// TIA Portal project "Proyecto_final" (V15.1)

(* hardware
DEVICE "S71500/ET200MP station_1"  S7-1500 station
   slot 0: "Rail_0"  Rack  6ES7 590-1***0-0AA0
   slot 1: "PLC_1"  CPU 1516-3 PN/DP  6ES7 516-3AN01-0AB0  V2.6
      slot 3: "CPU display_1"  6ES7591-1BA00-0AA0
   slot 2: "AI 8xU/I/RTD/TC ST_1"  AI 8xU/I/RTD/TC ST  6ES7 531-7KF00-0AB0  V2.2
   slot 3: "AQ 4xU/I ST_1"  AQ 4xU/I ST  6ES7 532-5HD00-0AB0  V2.2
   slot 4: "DI 32x24VDC HF_1"  DI 32x24VDC HF  6ES7 521-1BL00-0AB0  V2.1
   slot 5: "DQ 32x24VDC/0.5A HF_1"  DQ 32x24VDC/0.5A HF  6ES7 522-1BL01-0AB0  V1.1
DEVICE "S7-1200 station_1"  S7-1200 Station
   slot 0: "Rack_0"  S7-1200 Rack  Rack  V1.0
   slot 1: "PLC_2"  CPU 1215C DC/DC/DC  6ES7 215-1AG40-0XB0  V4.2
DEVICE "S7-1200 station_2"  S7-1200 Station
   slot 0: "Rack_0"  S7-1200 Rack  Rack  V1.0
   slot 1: "PLC_3"  CPU 1215C DC/DC/DC  6ES7 215-1AG40-0XB0  V4.2
DEVICE "HMI_1"  KTP400 Basic PN
   slot 0: "HMI_1"  KTP400 Basic PN  6AV2 123-2DB03-0AX0  15.1.0.0
   slot 1: "HMI_RT_1"  KTP400 Basic PN  6AV2 123-2DB03-0AX0  15.1.0.0
   slot 5: "HMI_1.IE_CP_1"  PROFINET Interface  15.0.1.0
      slot 1: "PROFINET Interface_1"  PROFINET Interface
         slot 1: "Port_1"  Port
DEVICE "HMI_2"  KTP400 Basic PN
   slot 0: "HMI_2"  KTP400 Basic PN  6AV2 123-2DB03-0AX0  15.1.0.0
   slot 1: "HMI_RT_2"  KTP400 Basic PN  6AV2 123-2DB03-0AX0  15.1.0.0
   slot 5: "HMI_2.IE_CP_1"  PROFINET Interface  15.0.1.0
      slot 1: "PROFINET Interface_1"  PROFINET Interface
         slot 1: "Port_1"  Port
DEVICE "HMI_3"  KTP400 Basic PN
   slot 0: "HMI_3"  KTP400 Basic PN  6AV2 123-2DB03-0AX0  15.1.0.0
   slot 1: "HMI_RT_3"  KTP400 Basic PN  6AV2 123-2DB03-0AX0  15.1.0.0
   slot 5: "HMI_3.IE_CP_1"  PROFINET Interface  15.0.1.0
      slot 1: "PROFINET Interface_1"  PROFINET Interface
         slot 1: "Port_1"  Port
DEVICE "SCALANCE X005"  SCALANCE X-Station
   slot 0: "SCALANCE X rack"  Rail
   slot 0: "Switch_1"  6GK5 005-0BA00-1AB2  V1.0
*)

// ===== PLC "PLC_1"  CPU 1516-3 PN/DP =====

VAR_GLOBAL   // PLC tag table "Default tag table"
   "Encendido" AT %M8.0 : Bool;
   "PE" AT %I17.3 : Bool;
   "Tag_1" AT %Q9.3 : Bool;
   "Tag_2" AT %Q9.4 : Bool;
   "LED_estado" AT %Q9.5 : Bool;
   "LED_PE" AT %Q9.6 : Bool;
   "Tag_3" AT %I17.4 : Bool;
   "Tag_4" AT %I17.5 : Bool;
   "Tag_5" AT %I17.6 : Bool;
END_VAR

DATA_BLOCK "PLC1_Ban"   // DB2
{ S7_Optimized_Access := 'FALSE' }
VERSION : 0.1
   VAR
      Ban_estado : Bool;
      Ban_dirección : UInt;
   END_VAR
BEGIN
END_DATA_BLOCK

// folder: System blocks/Program resources

DATA_BLOCK "IEC_Timer_0_DB"   // DB1
{ S7_Optimized_Access := 'TRUE' }
AUTHOR : Simatic
FAMILY : IEC
NAME : IEC_TMR
VERSION : 1.0
// stored: InstanceOfName IEC_TIMER
"IEC_TIMER"
BEGIN
END_DATA_BLOCK

// folder: (top level)

ORGANIZATION_BLOCK "Main"   // OB1, LAD, ProgramCycle
TITLE = Control de banda transportadora
{ S7_Optimized_Access := 'TRUE' }
VERSION : 0.1
   VAR_INPUT
      Initial_Call : Bool;   // Initial call of this OB
      Remanence : Bool;   // =True, if remanent data are available
   END_VAR
   VAR_TEMP   // added for the SCL form of the ladder/FBD networks
      _w1 : Bool;
   END_VAR
BEGIN

REGION Network 1: Control motor
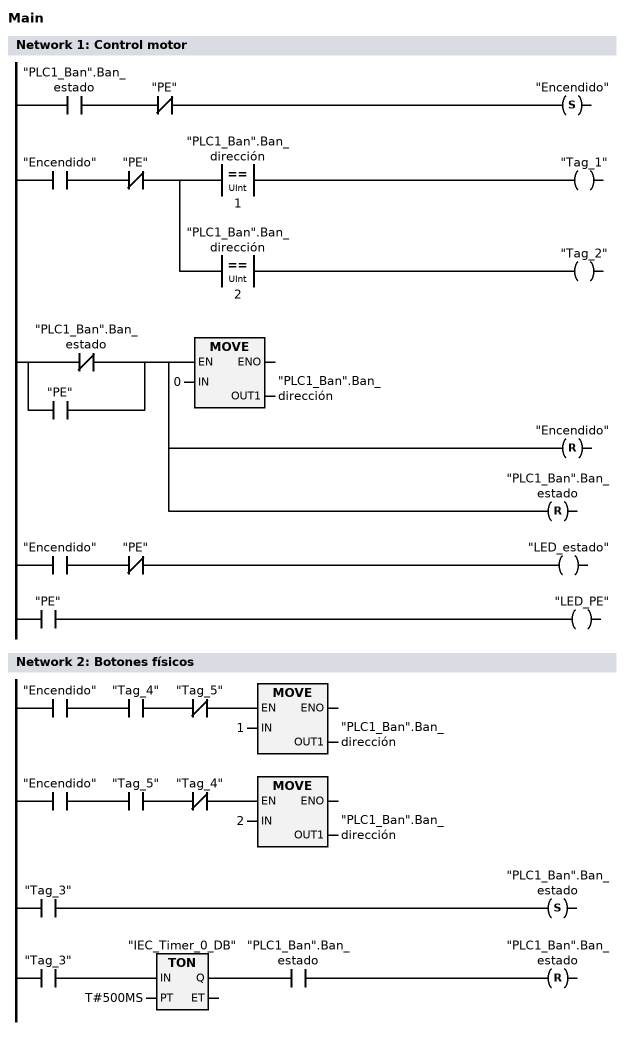
   RUNG wire#powerrail
      Contact( "PLC1_Ban".Ban_estado )
      I_Contact( "PE" )
      S_Coil( "Encendido" )
   END_RUNG
   RUNG wire#powerrail
      Contact( "Encendido" )
      I_Contact( "PE" )
      wire#w1
      { S7_Templates := "SrcType := UInt" } EQ_Contact(in1 := "PLC1_Ban".Ban_dirección, in2 := 1)
      Coil( "Tag_1" )
   END_RUNG
   RUNG wire#w1
      { S7_Templates := "SrcType := UInt" } EQ_Contact(in1 := "PLC1_Ban".Ban_dirección, in2 := 2)
      Coil( "Tag_2" )
   END_RUNG
   RUNG wire#powerrail
      I_Contact( "PLC1_Ban".Ban_estado )
      wire#w2
      Move(in := 0, out1 => "PLC1_Ban".Ban_dirección)
   END_RUNG
   RUNG wire#powerrail
      Contact( "PE" )
   END_RUNG wire#w2
   RUNG wire#w2
      R_Coil( "Encendido" )
   END_RUNG
   RUNG wire#w2
      R_Coil( "PLC1_Ban".Ban_estado )
   END_RUNG
   RUNG wire#powerrail
      Contact( "Encendido" )
      I_Contact( "PE" )
      Coil( "LED_estado" )
   END_RUNG
   RUNG wire#powerrail
      Contact( "PE" )
      Coil( "LED_PE" )
   END_RUNG
   // the same network as SCL:
   IF "PLC1_Ban".Ban_estado AND NOT "PE" THEN "Encendido" := TRUE; END_IF;
   #_w1 := "Encendido" AND NOT "PE";
   "Tag_1" := #_w1 AND ("PLC1_Ban".Ban_dirección = 1);
   "Tag_2" := #_w1 AND ("PLC1_Ban".Ban_dirección = 2);
   IF NOT "PLC1_Ban".Ban_estado OR "PE" THEN
       "PLC1_Ban".Ban_dirección := 0;
       "Encendido" := FALSE;
       "PLC1_Ban".Ban_estado := FALSE;
   END_IF;
   "LED_estado" := "Encendido" AND NOT "PE";
   "LED_PE" := "PE";
END_REGION

REGION Network 2: Botones físicos
   IF "Encendido" AND "Tag_4" AND NOT "Tag_5" THEN "PLC1_Ban".Ban_dirección := 1; END_IF;
   IF "Encendido" AND "Tag_5" AND NOT "Tag_4" THEN "PLC1_Ban".Ban_dirección := 2; END_IF;
   IF "Tag_3" THEN "PLC1_Ban".Ban_estado := TRUE; END_IF;
   "IEC_Timer_0_DB".TON(IN := "Tag_3", PT := T#500MS);
   IF "IEC_Timer_0_DB".Q AND "PLC1_Ban".Ban_estado THEN "PLC1_Ban".Ban_estado := FALSE; END_IF;
END_REGION
END_ORGANIZATION_BLOCK

// ===== PLC "PLC_2"  CPU 1215C DC/DC/DC =====

VAR_GLOBAL   // PLC tag table "Default tag table"
   "Rev_Detección" AT %M0.1 : Bool;
   "Rev_especial" AT %MW4 : UInt;
   "Rev_estado" AT %M0.0 : Bool;
   "Rev_progreso" AT %MW2 : Int;
   "B4" AT %I0.0 : Bool;
   "F3" AT %Q0.0 : Bool;
   "F2" AT %Q0.1 : Bool;
   "F1" AT %Q0.2 : Bool;
   "Piston_arriba" AT %Q0.3 : Bool;
   "Piston_abajo" AT %Q0.4 : Bool;
   "PE" AT %I0.4 : Bool;
   "Sens_abajo" AT %I0.5 : Bool;
   "Sens_arriba" AT %I0.6 : Bool;
   "B3" AT %I0.1 : Bool;
   "B2" AT %I0.2 : Bool;
   "B1" AT %I0.3 : Bool;
   "Encendido" AT %M0.2 : Bool;
   "Fin" AT %M0.3 : Bool;
   "Ciclo" AT %M0.4 : Bool;
   "Mem_pos" AT %M0.5 : Bool;
   "Cuenta_add" AT %MW6 : Int;
   "Reset" AT %M0.6 : Bool;
   "Skip" AT %M0.7 : Bool;
   "Tag_1" AT %M8.0 : Bool;
END_VAR

DATA_BLOCK "PLC2_Rev"   // DB5
{ S7_Optimized_Access := 'FALSE' }
VERSION : 0.1
   VAR
      Rev_Detección : Bool;
      Rev_especial : UInt;
      Rev_estado : Bool;
      Rev_progreso : Int;
   END_VAR
BEGIN
END_DATA_BLOCK

// folder: System blocks/Program resources

DATA_BLOCK "IEC_Timer_0_DB"   // DB1
{ S7_Optimized_Access := 'TRUE' }
AUTHOR : Simatic
FAMILY : IEC
NAME : IEC_TMR
VERSION : 1.0
// stored: InstanceOfName IEC_TIMER
"IEC_TIMER"
BEGIN
END_DATA_BLOCK

DATA_BLOCK "IEC_Counter_0_DB"   // DB2
{ S7_Optimized_Access := 'TRUE' }
AUTHOR : Simatic
FAMILY : IEC
NAME : CNTR
VERSION : 1.0
// stored: InstanceOfName IEC_COUNTER
"IEC_COUNTER"
BEGIN
END_DATA_BLOCK

DATA_BLOCK "IEC_Timer_0_DB_2"   // DB3
{ S7_Optimized_Access := 'TRUE' }
AUTHOR : Simatic
FAMILY : IEC
NAME : IEC_TMR
VERSION : 1.0
// stored: InstanceOfName IEC_TIMER
"IEC_TIMER"
BEGIN
END_DATA_BLOCK

DATA_BLOCK "IEC_Timer_0_DB_1"   // DB4
{ S7_Optimized_Access := 'TRUE' }
AUTHOR : Simatic
FAMILY : IEC
NAME : IEC_TMR
VERSION : 1.0
// stored: InstanceOfName IEC_TIMER
"IEC_TIMER"
BEGIN
END_DATA_BLOCK

DATA_BLOCK "IEC_Timer_0_DB_3"   // DB6
{ S7_Optimized_Access := 'TRUE' }
AUTHOR : Simatic
FAMILY : IEC
NAME : IEC_TMR
VERSION : 1.0
// stored: InstanceOfName IEC_TIMER
"IEC_TIMER"
BEGIN
END_DATA_BLOCK

DATA_BLOCK "IEC_Timer_0_DB_4"   // DB7
{ S7_Optimized_Access := 'TRUE' }
AUTHOR : Simatic
FAMILY : IEC
NAME : IEC_TMR
VERSION : 1.0
// stored: InstanceOfName IEC_TIMER
"IEC_TIMER"
BEGIN
END_DATA_BLOCK

DATA_BLOCK "IEC_Timer_0_DB_5"   // DB8
{ S7_Optimized_Access := 'TRUE' }
AUTHOR : Simatic
FAMILY : IEC
NAME : IEC_TMR
VERSION : 1.0
// stored: InstanceOfName IEC_TIMER
"IEC_TIMER"
BEGIN
END_DATA_BLOCK

// folder: (top level)

ORGANIZATION_BLOCK "Main"   // OB1, LAD, ProgramCycle
TITLE = Revolvedora
{ S7_Optimized_Access := 'TRUE' }
VERSION : 0.1
   VAR_INPUT
      Initial_Call : Bool;   // Initial call of this OB
      Remanence : Bool;   // =True, if remanent data are available
   END_VAR
   VAR_TEMP   // added for the SCL form of the ladder/FBD networks
      _w1 : Bool;
   END_VAR
BEGIN

REGION Network 1
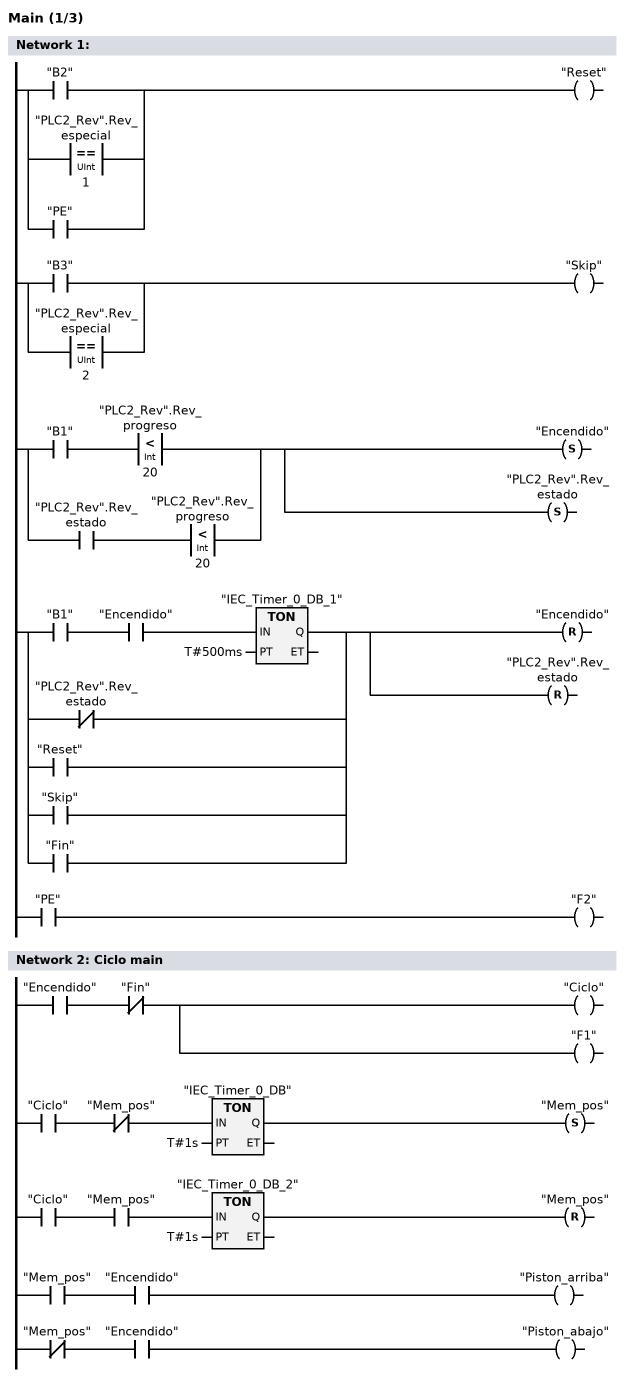
   "Reset" := "B2" OR ("PLC2_Rev".Rev_especial = 1) OR "PE";
   "Skip" := "B3" OR ("PLC2_Rev".Rev_especial = 2);
   IF ("B1" AND ("PLC2_Rev".Rev_progreso < 20)) OR ("PLC2_Rev".Rev_estado AND ("PLC2_Rev".Rev_progreso < 20)) THEN
       "Encendido" := TRUE;
       "PLC2_Rev".Rev_estado := TRUE;
   END_IF;
   "IEC_Timer_0_DB_1".TON(IN := "B1" AND "Encendido", PT := T#500ms);
   IF "IEC_Timer_0_DB_1".Q OR NOT "PLC2_Rev".Rev_estado OR "Reset" OR "Skip" OR "Fin" THEN
       "Encendido" := FALSE;
       "PLC2_Rev".Rev_estado := FALSE;
   END_IF;
   "F2" := "PE";
END_REGION

REGION Network 2: Ciclo main
   "Ciclo" := "Encendido" AND NOT "Fin";
   "F1" := "Ciclo";
   "IEC_Timer_0_DB".TON(IN := "Ciclo" AND NOT "Mem_pos", PT := T#1s);
   IF "IEC_Timer_0_DB".Q THEN "Mem_pos" := TRUE; END_IF;
   "IEC_Timer_0_DB_2".TON(IN := "Ciclo" AND "Mem_pos", PT := T#1s);
   IF "IEC_Timer_0_DB_2".Q THEN "Mem_pos" := FALSE; END_IF;
   "Piston_arriba" := "Mem_pos" AND "Encendido";
   "Piston_abajo" := NOT "Mem_pos" AND "Encendido";
END_REGION

REGION Network 3: Fin
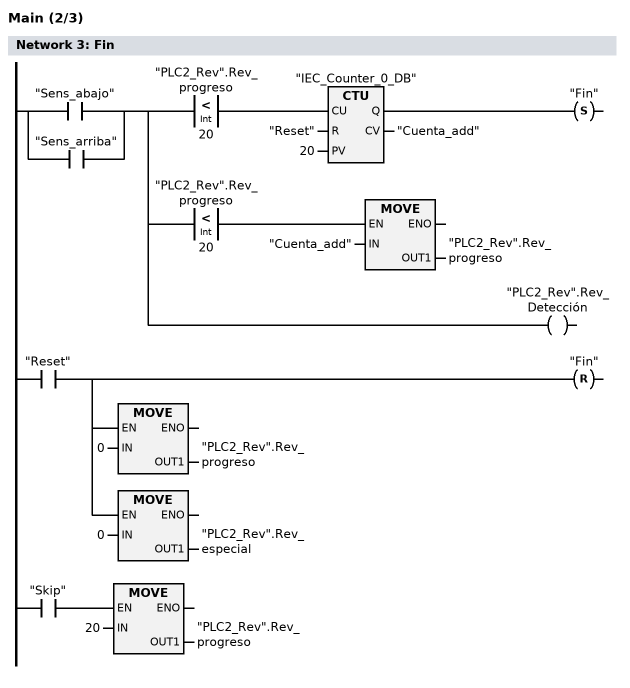
   #_w1 := "Sens_abajo" OR "Sens_arriba";
   "IEC_Counter_0_DB".CTU(CU := #_w1 AND ("PLC2_Rev".Rev_progreso < 20),
                          R := "Reset",
                          PV := 20,
                          CV => "Cuenta_add");
   IF "IEC_Counter_0_DB".Q THEN "Fin" := TRUE; END_IF;
   IF #_w1 AND ("PLC2_Rev".Rev_progreso < 20) THEN "PLC2_Rev".Rev_progreso := "Cuenta_add"; END_IF;
   "PLC2_Rev".Rev_Detección := #_w1;
   IF "Reset" THEN
       "Fin" := FALSE;
       "PLC2_Rev".Rev_progreso := 0;
       "PLC2_Rev".Rev_especial := 0;
   END_IF;
   IF "Skip" THEN "PLC2_Rev".Rev_progreso := 20; END_IF;
END_REGION

REGION Network 4: DB_control
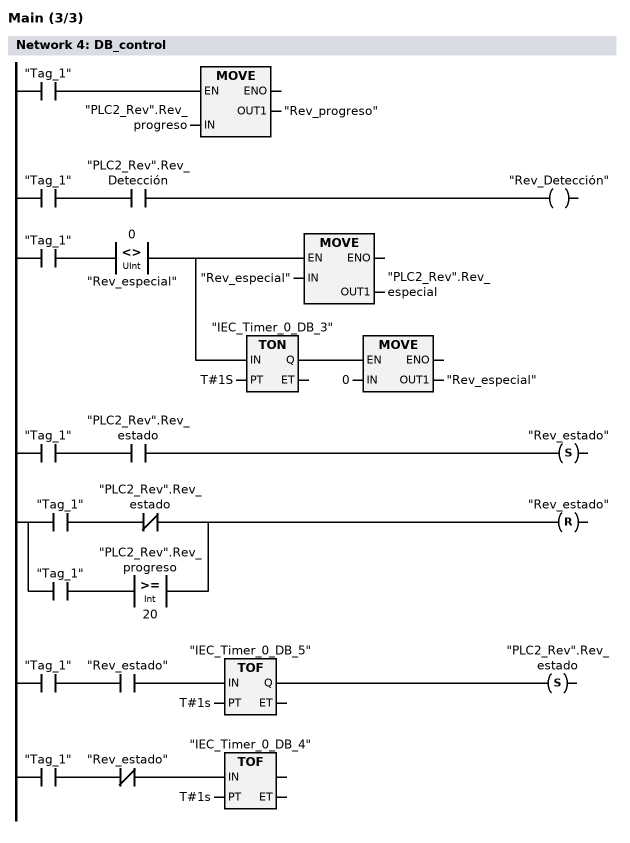
   IF "Tag_1" THEN "Rev_progreso" := "PLC2_Rev".Rev_progreso; END_IF;
   "Rev_Detección" := "Tag_1" AND "PLC2_Rev".Rev_Detección;
   #_w1 := "Tag_1" AND (0 <> "Rev_especial");
   IF #_w1 THEN "PLC2_Rev".Rev_especial := "Rev_especial"; END_IF;
   "IEC_Timer_0_DB_3".TON(IN := #_w1, PT := T#1S);
   IF "IEC_Timer_0_DB_3".Q THEN "Rev_especial" := 0; END_IF;
   IF "Tag_1" AND "PLC2_Rev".Rev_estado THEN "Rev_estado" := TRUE; END_IF;
   IF ("Tag_1" AND NOT "PLC2_Rev".Rev_estado) OR ("Tag_1" AND ("PLC2_Rev".Rev_progreso >= 20)) THEN
       "Rev_estado" := FALSE;
   END_IF;
   "IEC_Timer_0_DB_5".TOF(IN := "Tag_1" AND "Rev_estado", PT := T#1s);
   IF "IEC_Timer_0_DB_5".Q THEN "PLC2_Rev".Rev_estado := TRUE; END_IF;
   "IEC_Timer_0_DB_4".TOF(IN := "Tag_1" AND NOT "Rev_estado", PT := T#1s);
END_REGION
END_ORGANIZATION_BLOCK

// ===== PLC "PLC_3"  CPU 1215C DC/DC/DC =====

VAR_GLOBAL   // PLC tag table "Default tag table"
   "Emp_Estado" AT %M4.0 : Bool;
   "Emp_Especial" AT %MW0 : UInt;
   "Emp_Detección" AT %M4.1 : Bool;
   "Emp_Progreso" AT %MW2 : Int;
   "Start" AT %I1.3 : Bool;
   "Reiniciar" AT %I1.4 : Bool;
   "Skip" AT %I1.5 : Bool;
   "Encendido" AT %M4.2 : Bool;
   "Motor" AT %Q0.2 : Bool;
   "Fin" AT %M4.3 : Bool;
   "Reset" AT %M4.4 : Bool;
   "Detector" AT %I0.0 : Bool;
   "Emp_progreso_trans" AT %MW5 : Int;
END_VAR

DATA_BLOCK "PLC3_emp"   // DB3
{ S7_Optimized_Access := 'FALSE' }
VERSION : 0.1
   VAR
      Emp_estado : Bool;
      Emp_especial : UInt;
      Emp_detección : Bool;
      Emp_progreso : Int;
   END_VAR
BEGIN
END_DATA_BLOCK

// folder: System blocks/Program resources

DATA_BLOCK "IEC_Timer_0_DB"   // DB1
{ S7_Optimized_Access := 'TRUE' }
AUTHOR : Simatic
FAMILY : IEC
NAME : IEC_TMR
VERSION : 1.0
// stored: InstanceOfName IEC_TIMER
"IEC_TIMER"
BEGIN
END_DATA_BLOCK

DATA_BLOCK "IEC_Counter_0_DB"   // DB2
{ S7_Optimized_Access := 'TRUE' }
AUTHOR : Simatic
FAMILY : IEC
NAME : CNTR
VERSION : 1.0
// stored: InstanceOfName IEC_COUNTER
"IEC_COUNTER"
BEGIN
END_DATA_BLOCK

DATA_BLOCK "IEC_Timer_0_DB_1"   // DB4
{ S7_Optimized_Access := 'TRUE' }
AUTHOR : Simatic
FAMILY : IEC
NAME : IEC_TMR
VERSION : 1.0
// stored: InstanceOfName IEC_TIMER
"IEC_TIMER"
BEGIN
END_DATA_BLOCK

// folder: (top level)

ORGANIZATION_BLOCK "Main"   // OB1, LAD, ProgramCycle
TITLE = Empacadora circular
{ S7_Optimized_Access := 'TRUE' }
VERSION : 0.1
   VAR_INPUT
      Initial_Call : Bool;   // Initial call of this OB
      Remanence : Bool;   // =True, if remanent data are available
   END_VAR
BEGIN

REGION Network 1: Control Motor
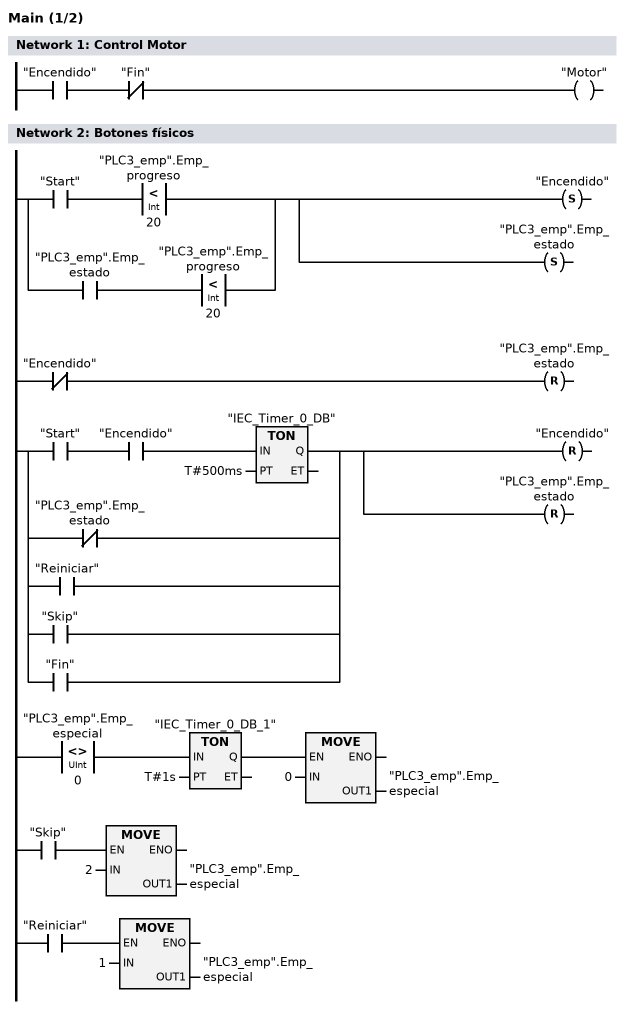
   RUNG wire#powerrail
      Contact( "Encendido" )
      I_Contact( "Fin" )
      Coil( "Motor" )
   END_RUNG
   // the same network as SCL:
   "Motor" := "Encendido" AND NOT "Fin";
END_REGION

REGION Network 2: Botones físicos
   IF ("Start" AND ("PLC3_emp".Emp_progreso < 20)) OR ("PLC3_emp".Emp_estado AND ("PLC3_emp".Emp_progreso < 20)) THEN
       "Encendido" := TRUE;
       "PLC3_emp".Emp_estado := TRUE;
   END_IF;
   IF NOT "Encendido" THEN "PLC3_emp".Emp_estado := FALSE; END_IF;
   "IEC_Timer_0_DB".TON(IN := "Start" AND "Encendido", PT := T#500ms);
   IF "IEC_Timer_0_DB".Q OR NOT "PLC3_emp".Emp_estado OR "Reiniciar" OR "Skip" OR "Fin" THEN
       "Encendido" := FALSE;
       "PLC3_emp".Emp_estado := FALSE;
   END_IF;
   "IEC_Timer_0_DB_1".TON(IN := "PLC3_emp".Emp_especial <> 0, PT := T#1s);
   IF "IEC_Timer_0_DB_1".Q THEN "PLC3_emp".Emp_especial := 0; END_IF;
   IF "Skip" THEN "PLC3_emp".Emp_especial := 2; END_IF;
   IF "Reiniciar" THEN "PLC3_emp".Emp_especial := 1; END_IF;
END_REGION

REGION Network 3: Cuenta
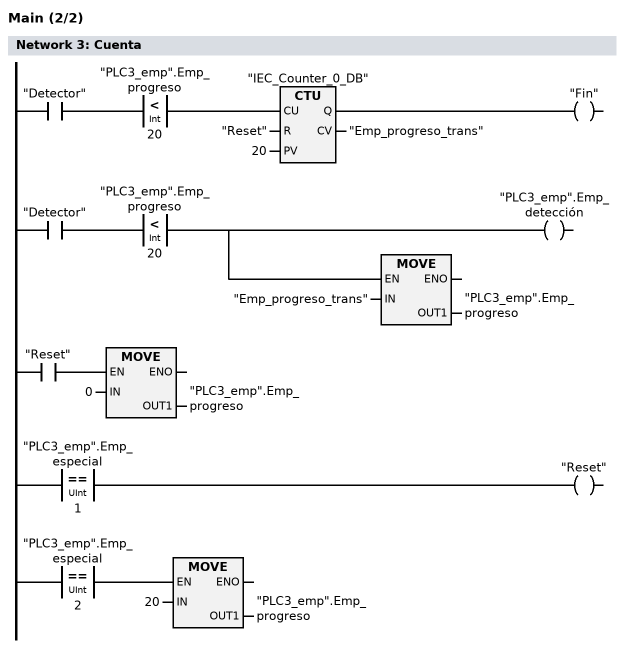
   "IEC_Counter_0_DB".CTU(CU := "Detector" AND ("PLC3_emp".Emp_progreso < 20),
                          R := "Reset",
                          PV := 20,
                          CV => "Emp_progreso_trans");
   "Fin" := "IEC_Counter_0_DB".Q;
   "PLC3_emp".Emp_detección := "Detector" AND ("PLC3_emp".Emp_progreso < 20);
   IF "PLC3_emp".Emp_detección THEN "PLC3_emp".Emp_progreso := "Emp_progreso_trans"; END_IF;
   IF "Reset" THEN "PLC3_emp".Emp_progreso := 0; END_IF;
   "Reset" := "PLC3_emp".Emp_especial = 1;
   IF "PLC3_emp".Emp_especial = 2 THEN "PLC3_emp".Emp_progreso := 20; END_IF;
END_REGION
END_ORGANIZATION_BLOCK

(* ===== HMI "HMI_RT_1" =====
system functions are stored by id; their names below are inferred from use
connection "Connection_1": ETHERNET, SMART_S7_1200_OMS
connection "HMI_Connection_1": ETHERNET, SMART_S7_1500_OMS

HMI tags "Default tag table"
   "Tag_ScreenNumber" : UInt, internal
   "Estado" : Bool = PLC PLC1_Ban.Ban_estado AT %DB2.DBX0.0, 500 ms
   "Dirección" : UInt = PLC PLC1_Ban.Ban_dirección AT %DB2.DBW2, 500 ms

text list "Estado": 0..1 'Apagado'; 1 'Encendido'

text list "Dirección": 0..1 'Apagado'; 1 'Adelante'; 2 'Reversa'

Template "Template_1" 480x272
   Button "Exit" at 388,227 size 63x44; TextOff 'Exit'; PictureOff "ExitRuntime_KTP400_Basic_PN_TR"; PictureOn "ExitRuntime_KTP400_Basic_PN_TR"
      on Release: StopRuntime(0)
   GraphicView "Logo" at 0,0 size 160x45; Picture "Logo of HMI_1"

screen "Banda transportadora" 480x272
   TextField "Text field_2" at 89,81 size 79x28; Text 'Estado:'
   TextField "Text field_3" at 61,129 size 107x28; Text 'Dirección:'
   Button "Button_2" at 214,193 size 96x55; TextOff 'Adelante'
      on Click: SetTag("Dirección", 1)
   Button "Button_3" at 348,192 size 96x55; TextOff 'Reversa'
      on Click: SetTag("Dirección", 2)
   GraphicView "Graphic view_1" at 0,3 size 176x48; Picture "Logo of HMI_1"
   TextField "Text field_6" at 179,6 size 265x33; Text 'Banda transportadora'
   Switch "Switch_1" at 22,196 size 147x51; CaptionText 'Switch'; TextOff 'Apagado'; TextOn 'Encendio'
      ProcessValue <- "Estado"
      on SwitchOff: SetTag("Estado", 0)
      on SwitchOn: SetTag("Estado", 1)
   SymbolicIOField "Symbolic I/O field_1" at 198,72 size 155x46; TextOff '0'; TextOn '1'; TextList "Estado"
      ProcessValue <- "Estado"
   SymbolicIOField "Symbolic I/O field_2" at 198,121 size 155x46; TextOn '1'; TextOff '0'; TextList "Dirección"
      ProcessValue <- "Dirección"
*)

(* ===== HMI "HMI_RT_2" =====
system functions are stored by id; their names below are inferred from use
connection "Connection_2": ETHERNET, SMART_S7_1200_OMS
connection "HMI_Connection_3": ETHERNET, SMART_S7_1200_OMS

HMI tags "Default tag table"
   "Tag_ScreenNumber" : UInt, internal
   "Detección" : Bool = PLC PLC2_Rev.Rev_Detección AT %DB5.DBX0.0, 100 ms
   "Especial" : UInt = PLC PLC2_Rev.Rev_especial AT %DB5.DBW2, 100 ms
   "Estado" : Bool = PLC PLC2_Rev.Rev_estado AT %DB5.DBX4.0, 100 ms
   "Progreso" : Int = PLC PLC2_Rev.Rev_progreso AT %DB5.DBW6, 100 ms

text list "Estado": 0..1 'Apagado'; 1 'Encendido'

text list "Dirección": 0..1 'Apagado'; 1 'Adelante'; 2 'Reversa'

Template "Template_1" 480x272
   GraphicView "Logo" at 0,0 size 160x45; Picture "Logo of HMI_2"

screen "Revolvedora" 480x272
   TextField "Text field_2" at 33,73 size 79x28; Text 'Estado:'
   TextField "Text field_3" at 0,133 size 112x28; Text 'Detección:'
   Button "Button_2" at 211,212 size 96x55; TextOff 'Reiniciar'
      on Click: SetTag("Estado", 0); SetTag("Especial", 1)
   Button "Button_3" at 348,212 size 96x55; TextOff 'Skip'
      on Click: SetTag("Estado", 0); SetTag("Especial", 2)
   GraphicView "Graphic view_1" at 0,3 size 176x48; Picture "Logo of HMI_1"
   TextField "Text field_6" at 179,6 size 154x33; Text 'Revolvedora'
   Switch "Switch_1" at 9,212 size 147x51; TextOn 'Encendio'; CaptionText 'Switch'; TextOff 'Apagado'
      on SwitchOff: SetTag("Estado", 0)
      on SwitchOn: SetTag("Estado", 1)
      ProcessValue <- "Estado"
   SymbolicIOField "Symbolic I/O field_1" at 120,64 size 155x46; TextOn '1'; TextOff '0'; TextList "Estado"
      ProcessValue <- "Estado"
   TextField "Text field_1" at 342,45 size 102x28; Text 'Progreso:'
   Bar "Bar_1" at 359,75 size 80x120; MinimumValue 0; MaximumValue 20
      ProcessValue <- "Progreso"
   Circle "Circle_1" at 176,123 size 48x48
      Appearance <- "Detección"
*)

(* ===== HMI "HMI_RT_3" =====
system functions are stored by id; their names below are inferred from use
connection "Connection_3": ETHERNET, SMART_S7_1200_OMS
connection "HMI_Connection_2": ETHERNET, SMART_S7_1200_OMS

HMI tags "Default tag table"
   "Tag_ScreenNumber" : UInt, internal
   "Estado" : Bool = PLC PLC3_emp.Emp_estado AT %DB3.DBX0.0, 100 ms
   "Especial" : UInt = PLC PLC3_emp.Emp_especial AT %DB3.DBW2, 100 ms
   "Detección" : Bool = PLC PLC3_emp.Emp_detección AT %DB3.DBX4.0, 100 ms
   "Progreso" : Int = PLC PLC3_emp.Emp_progreso AT %DB3.DBW6, 100 ms

text list "Estado": 0..1 'Apagado'; 1 'Encendido'

Template "Template_1" 480x272
   GraphicView "Logo" at 0,0 size 160x45; Picture "Logo of HMI_3"

screen "Empacadora" 480x272
   TextField "Text field_2" at 33,73 size 79x28; Text 'Estado:'
   TextField "Text field_3" at 0,133 size 112x28; Text 'Detección:'
   Button "Button_2" at 211,212 size 96x55; TextOff 'Reiniciar'
      on Click: SetTag("Estado", 0); SetTag("Especial", 1)
   Button "Button_3" at 348,212 size 96x55; TextOff 'Skip'
      on Click: SetTag("Estado", 0); SetTag("Especial", 2)
   GraphicView "Graphic view_1" at 0,3 size 176x48; Picture "Logo of HMI_1"
   TextField "Text field_6" at 179,6 size 153x33; Text 'Empacadora'
   Switch "Switch_1" at 9,212 size 147x51; TextOn 'Encendio'; CaptionText 'Switch'; TextOff 'Apagado'
      on SwitchOff: SetTag("Estado", 0)
      on SwitchOn: SetTag("Estado", 1)
      ProcessValue <- "Estado"
   SymbolicIOField "Symbolic I/O field_1" at 120,64 size 155x46; TextOn '1'; TextOff '0'; TextList "Estado"
      ProcessValue <- "Estado"
   TextField "Text field_1" at 342,45 size 102x28; Text 'Progreso:'
   Bar "Bar_1" at 359,75 size 80x120; MinimumValue 0; MaximumValue 20
      ProcessValue <- "Progreso"
   Circle "Circle_1" at 176,123 size 48x48
      Appearance <- "Detección"
*)